(* Logix 5000 project; controller FV vendor 1 type 14 code 217 rev 31.11; software revision 31.00; part 46 of 63 *)
(* tags used below, declared in another part *)
   CWD : CHECKWORD_FLAGS;
   Delphi_Does_Eng_Func : BOOL;
   FV_FV10C : PlantItem;   // FV10C
   FV_FV10J : PlantItem;   // FV10J
   FV_FV11C : PlantItem;   // FV11C
   FV_FV11J : PlantItem;   // FV11J
   FV_FV12C : PlantItem;   // FV12C
   FV_FV12J : PlantItem;   // FV12J
   FV_FV1C : PlantItem;   // FV1C
   FV_FV1J : PlantItem;   // FV1J
   FV_FV2C : PlantItem;   // FV2C
   FV_FV2J : PlantItem;   // FV2J
   FV_FV3C : PlantItem;   // FV3C
   FV_FV3J : PlantItem;   // FV3J
   FV_FV4C : PlantItem;   // FV4C
   FV_FV4J : PlantItem;   // FV4J
   FV_FV5C : PlantItem;   // FV5C
   FV_FV5J : PlantItem;   // FV5J
   FV_FV6C : PlantItem;   // FV6C
   FV_FV6J : PlantItem;   // FV6J
   FV_FV7C : PlantItem;   // FV7C
   FV_FV7J : PlantItem;   // FV7J
   FV_FV8C : PlantItem;   // FV8C
   FV_FV8J : PlantItem;   // FV8J
   FV_FV9C : PlantItem;   // FV9C
   FV_FV9J : PlantItem;   // FV9J
   FV_N255 : INT[255];   // Old Checkwords to keep Delphi working in the interim before full changeover.
(* FV_Common, continued *)

ROUTINE FV_Old_Checkword_Relaying   (* ladder *)
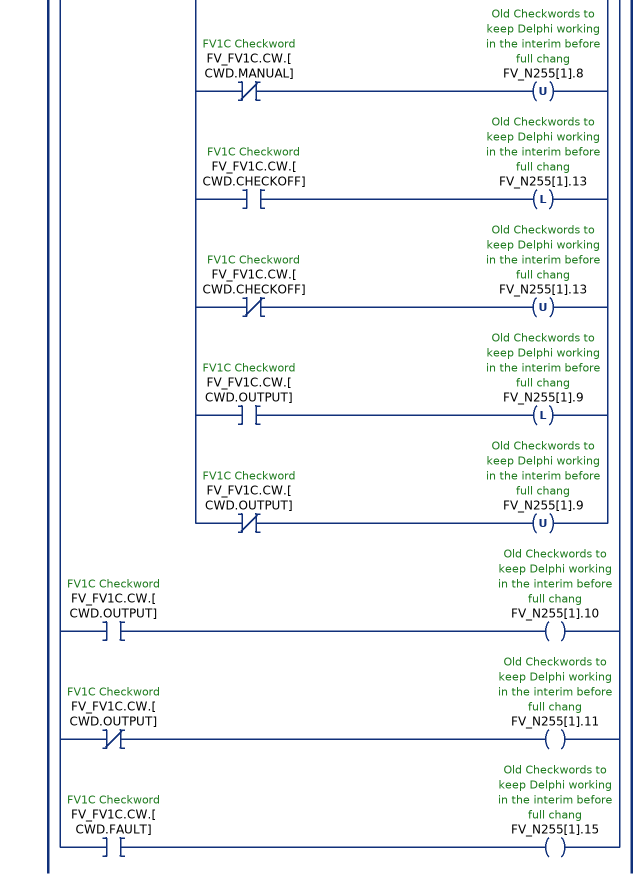
   0: [XIC(Delphi_Does_Eng_Func) [[XIC(FV_N255[1].8) [OTL(FV_FV1C.CW.[CWD.MANUAL]) ,XIC(FV_N255[1].9) OTL(FV_FV1C.CW.[CWD.MANDRV]) ,XIO(FV_N255[1].9) OTU(FV_FV1C.CW.[CWD.MANDRV]) ] ,XIO(FV_N255[1].8) [OTU(FV_FV1C.CW.[CWD.MANUAL]) ,[XIC(FV_FV1C.CW.[CWD.OUTPUT]) OTL(FV_N255[1].9) ,XIO(FV_FV1C.CW.[CWD.OUTPUT]) OTU(FV_N255[1].9) ] ] ] ,[XIC(FV_N255[1].13) OTL(FV_FV1C.CW.[CWD.CHECKOFF]) ,XIO(FV_N255[1].13) OTU(FV_FV1C.CW.[CWD.CHECKOFF]) ] ] ,XIO(Delphi_Does_Eng_Func) [[XIC(FV_FV1C.CW.[CWD.MANUAL]) OTL(FV_N255[1].8) ,XIO(FV_FV1C.CW.[CWD.MANUAL]) OTU(FV_N255[1].8) ] ,[XIC(FV_FV1C.CW.[CWD.CHECKOFF]) OTL(FV_N255[1].13) ,XIO(FV_FV1C.CW.[CWD.CHECKOFF]) OTU(FV_N255[1].13) ] ,[XIC(FV_FV1C.CW.[CWD.OUTPUT]) OTL(FV_N255[1].9) ,XIO(FV_FV1C.CW.[CWD.OUTPUT]) OTU(FV_N255[1].9) ] ] ,XIC(FV_FV1C.CW.[CWD.OUTPUT]) OTE(FV_N255[1].10) ,XIO(FV_FV1C.CW.[CWD.OUTPUT]) OTE(FV_N255[1].11) ,XIC(FV_FV1C.CW.[CWD.FAULT]) OTE(FV_N255[1].15) ];
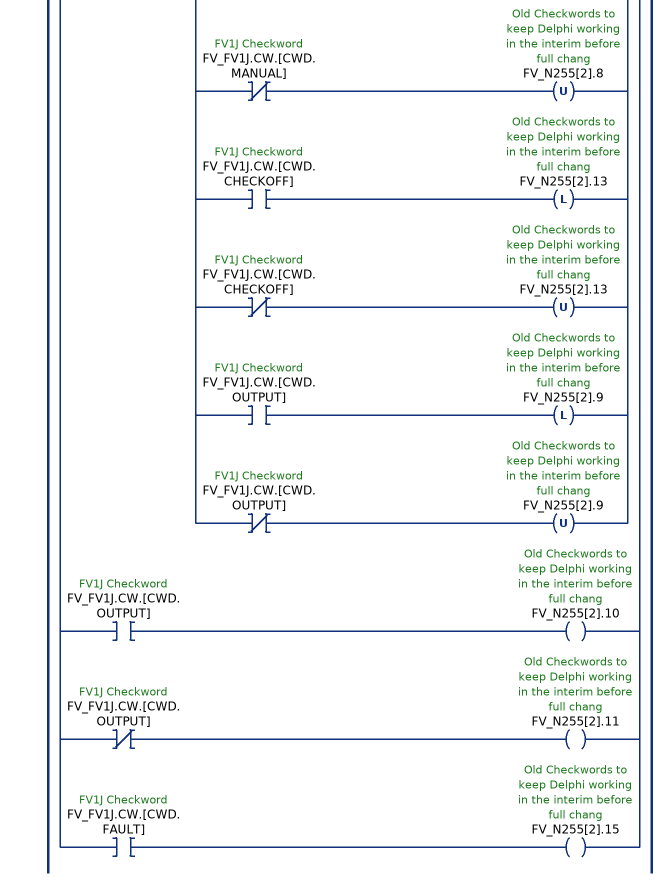
   1: [XIC(Delphi_Does_Eng_Func) [[XIC(FV_N255[2].8) [OTL(FV_FV1J.CW.[CWD.MANUAL]) ,XIC(FV_N255[2].9) OTL(FV_FV1J.CW.[CWD.MANDRV]) ,XIO(FV_N255[2].9) OTU(FV_FV1J.CW.[CWD.MANDRV]) ] ,XIO(FV_N255[2].8) [OTU(FV_FV1J.CW.[CWD.MANUAL]) ,[XIC(FV_FV1J.CW.[CWD.OUTPUT]) OTL(FV_N255[2].9) ,XIO(FV_FV1J.CW.[CWD.OUTPUT]) OTU(FV_N255[2].9) ] ] ] ,[XIC(FV_N255[2].13) OTL(FV_FV1J.CW.[CWD.CHECKOFF]) ,XIO(FV_N255[2].13) OTU(FV_FV1J.CW.[CWD.CHECKOFF]) ] ] ,XIO(Delphi_Does_Eng_Func) [[XIC(FV_FV1J.CW.[CWD.MANUAL]) OTL(FV_N255[2].8) ,XIO(FV_FV1J.CW.[CWD.MANUAL]) OTU(FV_N255[2].8) ] ,[XIC(FV_FV1J.CW.[CWD.CHECKOFF]) OTL(FV_N255[2].13) ,XIO(FV_FV1J.CW.[CWD.CHECKOFF]) OTU(FV_N255[2].13) ] ,[XIC(FV_FV1J.CW.[CWD.OUTPUT]) OTL(FV_N255[2].9) ,XIO(FV_FV1J.CW.[CWD.OUTPUT]) OTU(FV_N255[2].9) ] ] ,XIC(FV_FV1J.CW.[CWD.OUTPUT]) OTE(FV_N255[2].10) ,XIO(FV_FV1J.CW.[CWD.OUTPUT]) OTE(FV_N255[2].11) ,XIC(FV_FV1J.CW.[CWD.FAULT]) OTE(FV_N255[2].15) ];
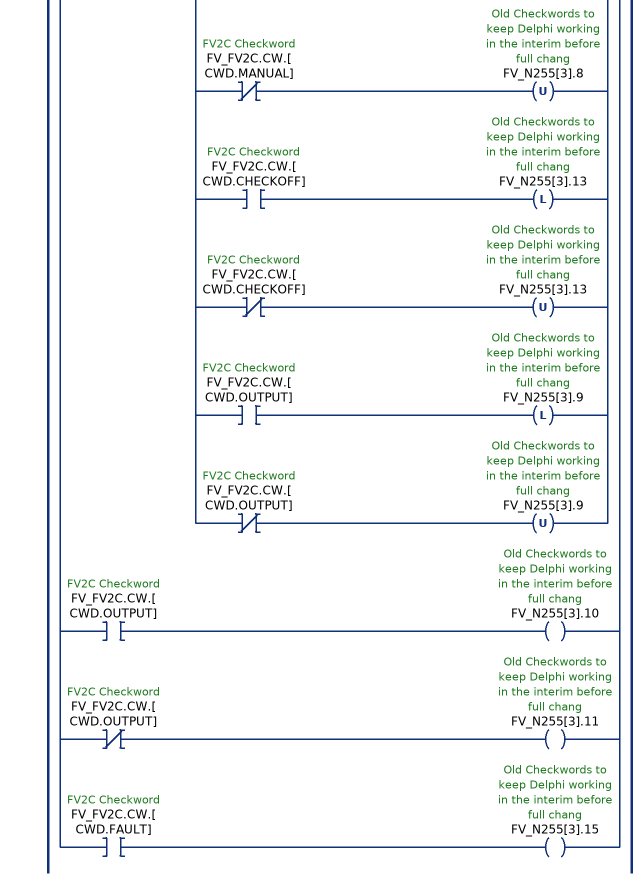
   2: [XIC(Delphi_Does_Eng_Func) [[XIC(FV_N255[3].8) [OTL(FV_FV2C.CW.[CWD.MANUAL]) ,XIC(FV_N255[3].9) OTL(FV_FV2C.CW.[CWD.MANDRV]) ,XIO(FV_N255[3].9) OTU(FV_FV2C.CW.[CWD.MANDRV]) ] ,XIO(FV_N255[3].8) [OTU(FV_FV2C.CW.[CWD.MANUAL]) ,[XIC(FV_FV2C.CW.[CWD.OUTPUT]) OTL(FV_N255[3].9) ,XIO(FV_FV2C.CW.[CWD.OUTPUT]) OTU(FV_N255[3].9) ] ] ] ,[XIC(FV_N255[3].13) OTL(FV_FV2C.CW.[CWD.CHECKOFF]) ,XIO(FV_N255[3].13) OTU(FV_FV2C.CW.[CWD.CHECKOFF]) ] ] ,XIO(Delphi_Does_Eng_Func) [[XIC(FV_FV2C.CW.[CWD.MANUAL]) OTL(FV_N255[3].8) ,XIO(FV_FV2C.CW.[CWD.MANUAL]) OTU(FV_N255[3].8) ] ,[XIC(FV_FV2C.CW.[CWD.CHECKOFF]) OTL(FV_N255[3].13) ,XIO(FV_FV2C.CW.[CWD.CHECKOFF]) OTU(FV_N255[3].13) ] ,[XIC(FV_FV2C.CW.[CWD.OUTPUT]) OTL(FV_N255[3].9) ,XIO(FV_FV2C.CW.[CWD.OUTPUT]) OTU(FV_N255[3].9) ] ] ,XIC(FV_FV2C.CW.[CWD.OUTPUT]) OTE(FV_N255[3].10) ,XIO(FV_FV2C.CW.[CWD.OUTPUT]) OTE(FV_N255[3].11) ,XIC(FV_FV2C.CW.[CWD.FAULT]) OTE(FV_N255[3].15) ];
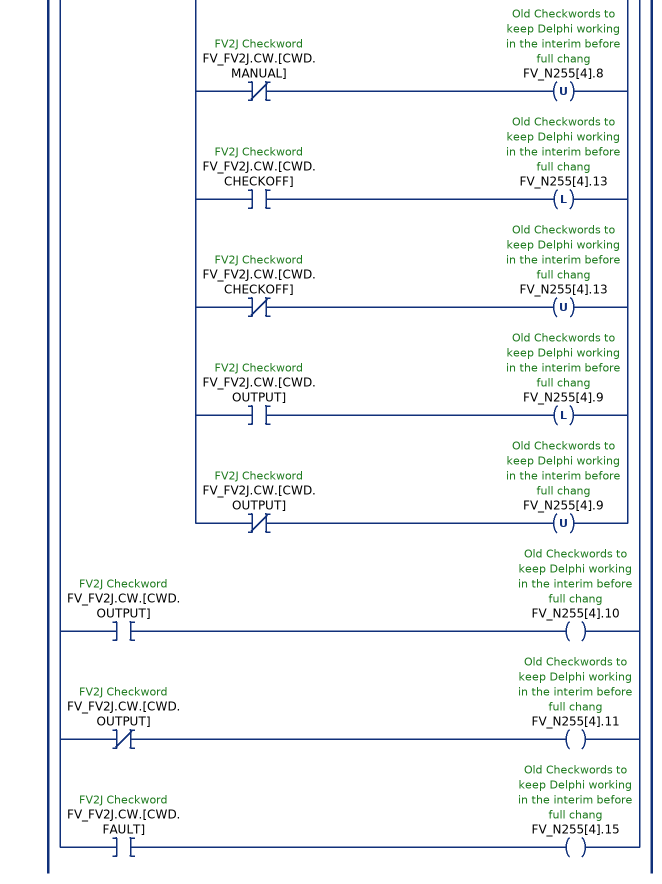
   3: [XIC(Delphi_Does_Eng_Func) [[XIC(FV_N255[4].8) [OTL(FV_FV2J.CW.[CWD.MANUAL]) ,XIC(FV_N255[4].9) OTL(FV_FV2J.CW.[CWD.MANDRV]) ,XIO(FV_N255[4].9) OTU(FV_FV2J.CW.[CWD.MANDRV]) ] ,XIO(FV_N255[4].8) [OTU(FV_FV2J.CW.[CWD.MANUAL]) ,[XIC(FV_FV2J.CW.[CWD.OUTPUT]) OTL(FV_N255[4].9) ,XIO(FV_FV2J.CW.[CWD.OUTPUT]) OTU(FV_N255[4].9) ] ] ] ,[XIC(FV_N255[4].13) OTL(FV_FV2J.CW.[CWD.CHECKOFF]) ,XIO(FV_N255[4].13) OTU(FV_FV2J.CW.[CWD.CHECKOFF]) ] ] ,XIO(Delphi_Does_Eng_Func) [[XIC(FV_FV2J.CW.[CWD.MANUAL]) OTL(FV_N255[4].8) ,XIO(FV_FV2J.CW.[CWD.MANUAL]) OTU(FV_N255[4].8) ] ,[XIC(FV_FV2J.CW.[CWD.CHECKOFF]) OTL(FV_N255[4].13) ,XIO(FV_FV2J.CW.[CWD.CHECKOFF]) OTU(FV_N255[4].13) ] ,[XIC(FV_FV2J.CW.[CWD.OUTPUT]) OTL(FV_N255[4].9) ,XIO(FV_FV2J.CW.[CWD.OUTPUT]) OTU(FV_N255[4].9) ] ] ,XIC(FV_FV2J.CW.[CWD.OUTPUT]) OTE(FV_N255[4].10) ,XIO(FV_FV2J.CW.[CWD.OUTPUT]) OTE(FV_N255[4].11) ,XIC(FV_FV2J.CW.[CWD.FAULT]) OTE(FV_N255[4].15) ];
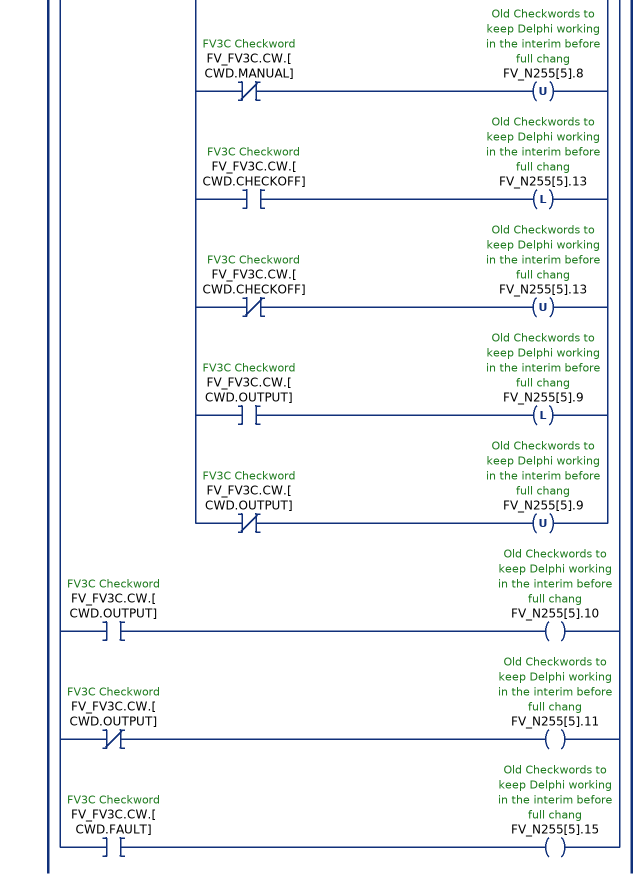
   4: [XIC(Delphi_Does_Eng_Func) [[XIC(FV_N255[5].8) [OTL(FV_FV3C.CW.[CWD.MANUAL]) ,XIC(FV_N255[5].9) OTL(FV_FV3C.CW.[CWD.MANDRV]) ,XIO(FV_N255[5].9) OTU(FV_FV3C.CW.[CWD.MANDRV]) ] ,XIO(FV_N255[5].8) [OTU(FV_FV3C.CW.[CWD.MANUAL]) ,[XIC(FV_FV3C.CW.[CWD.OUTPUT]) OTL(FV_N255[5].9) ,XIO(FV_FV3C.CW.[CWD.OUTPUT]) OTU(FV_N255[5].9) ] ] ] ,[XIC(FV_N255[5].13) OTL(FV_FV3C.CW.[CWD.CHECKOFF]) ,XIO(FV_N255[5].13) OTU(FV_FV3C.CW.[CWD.CHECKOFF]) ] ] ,XIO(Delphi_Does_Eng_Func) [[XIC(FV_FV3C.CW.[CWD.MANUAL]) OTL(FV_N255[5].8) ,XIO(FV_FV3C.CW.[CWD.MANUAL]) OTU(FV_N255[5].8) ] ,[XIC(FV_FV3C.CW.[CWD.CHECKOFF]) OTL(FV_N255[5].13) ,XIO(FV_FV3C.CW.[CWD.CHECKOFF]) OTU(FV_N255[5].13) ] ,[XIC(FV_FV3C.CW.[CWD.OUTPUT]) OTL(FV_N255[5].9) ,XIO(FV_FV3C.CW.[CWD.OUTPUT]) OTU(FV_N255[5].9) ] ] ,XIC(FV_FV3C.CW.[CWD.OUTPUT]) OTE(FV_N255[5].10) ,XIO(FV_FV3C.CW.[CWD.OUTPUT]) OTE(FV_N255[5].11) ,XIC(FV_FV3C.CW.[CWD.FAULT]) OTE(FV_N255[5].15) ];
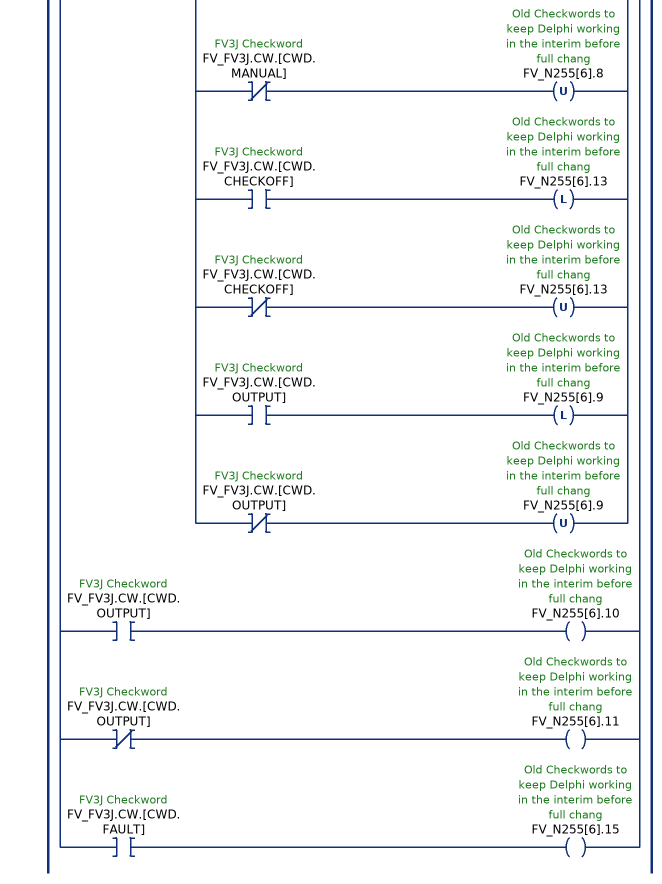
   5: [XIC(Delphi_Does_Eng_Func) [[XIC(FV_N255[6].8) [OTL(FV_FV3J.CW.[CWD.MANUAL]) ,XIC(FV_N255[6].9) OTL(FV_FV3J.CW.[CWD.MANDRV]) ,XIO(FV_N255[6].9) OTU(FV_FV3J.CW.[CWD.MANDRV]) ] ,XIO(FV_N255[6].8) [OTU(FV_FV3J.CW.[CWD.MANUAL]) ,[XIC(FV_FV3J.CW.[CWD.OUTPUT]) OTL(FV_N255[6].9) ,XIO(FV_FV3J.CW.[CWD.OUTPUT]) OTU(FV_N255[6].9) ] ] ] ,[XIC(FV_N255[6].13) OTL(FV_FV3J.CW.[CWD.CHECKOFF]) ,XIO(FV_N255[6].13) OTU(FV_FV3J.CW.[CWD.CHECKOFF]) ] ] ,XIO(Delphi_Does_Eng_Func) [[XIC(FV_FV3J.CW.[CWD.MANUAL]) OTL(FV_N255[6].8) ,XIO(FV_FV3J.CW.[CWD.MANUAL]) OTU(FV_N255[6].8) ] ,[XIC(FV_FV3J.CW.[CWD.CHECKOFF]) OTL(FV_N255[6].13) ,XIO(FV_FV3J.CW.[CWD.CHECKOFF]) OTU(FV_N255[6].13) ] ,[XIC(FV_FV3J.CW.[CWD.OUTPUT]) OTL(FV_N255[6].9) ,XIO(FV_FV3J.CW.[CWD.OUTPUT]) OTU(FV_N255[6].9) ] ] ,XIC(FV_FV3J.CW.[CWD.OUTPUT]) OTE(FV_N255[6].10) ,XIO(FV_FV3J.CW.[CWD.OUTPUT]) OTE(FV_N255[6].11) ,XIC(FV_FV3J.CW.[CWD.FAULT]) OTE(FV_N255[6].15) ];
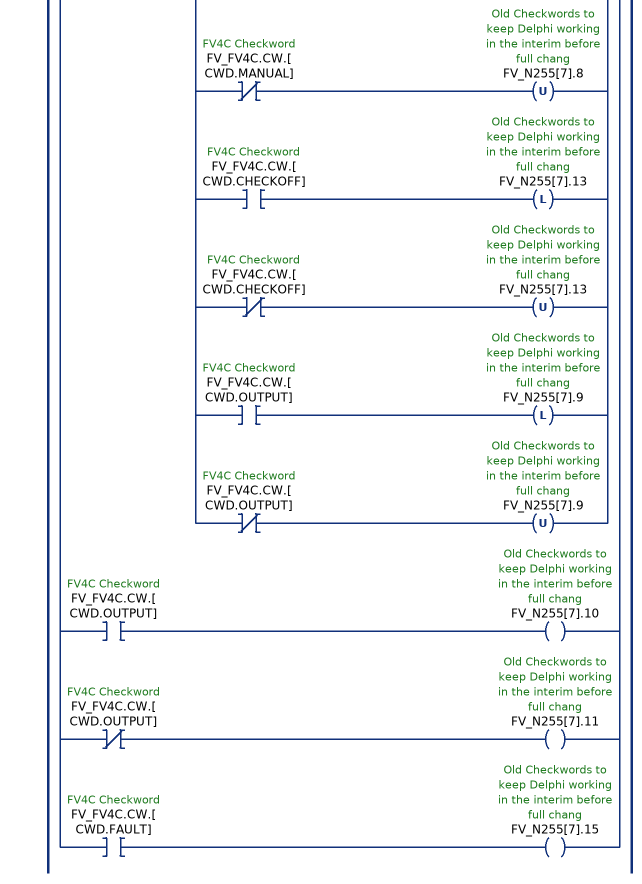
   6: [XIC(Delphi_Does_Eng_Func) [[XIC(FV_N255[7].8) [OTL(FV_FV4C.CW.[CWD.MANUAL]) ,XIC(FV_N255[7].9) OTL(FV_FV4C.CW.[CWD.MANDRV]) ,XIO(FV_N255[7].9) OTU(FV_FV4C.CW.[CWD.MANDRV]) ] ,XIO(FV_N255[7].8) [OTU(FV_FV4C.CW.[CWD.MANUAL]) ,[XIC(FV_FV4C.CW.[CWD.OUTPUT]) OTL(FV_N255[7].9) ,XIO(FV_FV4C.CW.[CWD.OUTPUT]) OTU(FV_N255[7].9) ] ] ] ,[XIC(FV_N255[7].13) OTL(FV_FV4C.CW.[CWD.CHECKOFF]) ,XIO(FV_N255[7].13) OTU(FV_FV4C.CW.[CWD.CHECKOFF]) ] ] ,XIO(Delphi_Does_Eng_Func) [[XIC(FV_FV4C.CW.[CWD.MANUAL]) OTL(FV_N255[7].8) ,XIO(FV_FV4C.CW.[CWD.MANUAL]) OTU(FV_N255[7].8) ] ,[XIC(FV_FV4C.CW.[CWD.CHECKOFF]) OTL(FV_N255[7].13) ,XIO(FV_FV4C.CW.[CWD.CHECKOFF]) OTU(FV_N255[7].13) ] ,[XIC(FV_FV4C.CW.[CWD.OUTPUT]) OTL(FV_N255[7].9) ,XIO(FV_FV4C.CW.[CWD.OUTPUT]) OTU(FV_N255[7].9) ] ] ,XIC(FV_FV4C.CW.[CWD.OUTPUT]) OTE(FV_N255[7].10) ,XIO(FV_FV4C.CW.[CWD.OUTPUT]) OTE(FV_N255[7].11) ,XIC(FV_FV4C.CW.[CWD.FAULT]) OTE(FV_N255[7].15) ];
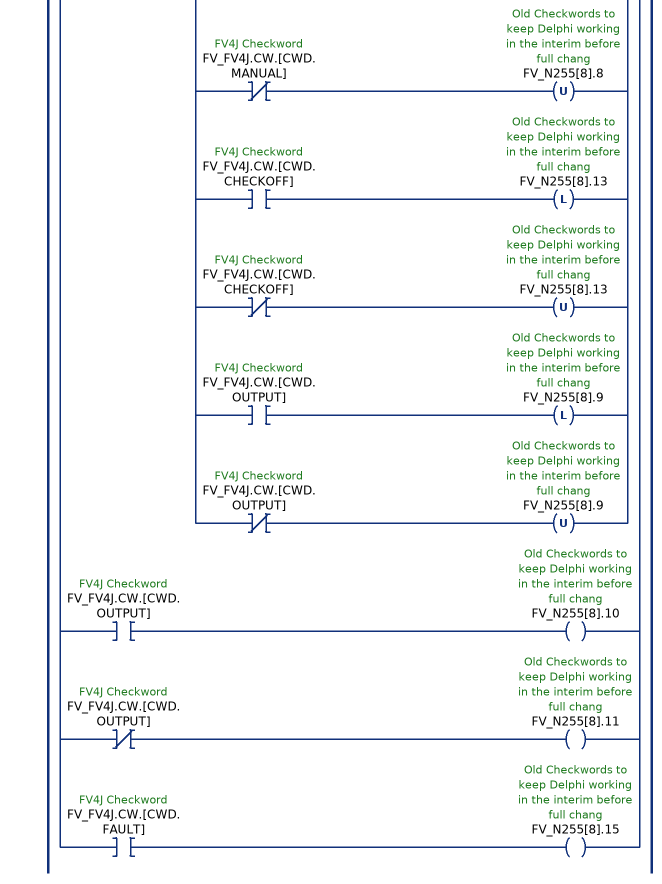
   7: [XIC(Delphi_Does_Eng_Func) [[XIC(FV_N255[8].8) [OTL(FV_FV4J.CW.[CWD.MANUAL]) ,XIC(FV_N255[8].9) OTL(FV_FV4J.CW.[CWD.MANDRV]) ,XIO(FV_N255[8].9) OTU(FV_FV4J.CW.[CWD.MANDRV]) ] ,XIO(FV_N255[8].8) [OTU(FV_FV4J.CW.[CWD.MANUAL]) ,[XIC(FV_FV4J.CW.[CWD.OUTPUT]) OTL(FV_N255[8].9) ,XIO(FV_FV4J.CW.[CWD.OUTPUT]) OTU(FV_N255[8].9) ] ] ] ,[XIC(FV_N255[8].13) OTL(FV_FV4J.CW.[CWD.CHECKOFF]) ,XIO(FV_N255[8].13) OTU(FV_FV4J.CW.[CWD.CHECKOFF]) ] ] ,XIO(Delphi_Does_Eng_Func) [[XIC(FV_FV4J.CW.[CWD.MANUAL]) OTL(FV_N255[8].8) ,XIO(FV_FV4J.CW.[CWD.MANUAL]) OTU(FV_N255[8].8) ] ,[XIC(FV_FV4J.CW.[CWD.CHECKOFF]) OTL(FV_N255[8].13) ,XIO(FV_FV4J.CW.[CWD.CHECKOFF]) OTU(FV_N255[8].13) ] ,[XIC(FV_FV4J.CW.[CWD.OUTPUT]) OTL(FV_N255[8].9) ,XIO(FV_FV4J.CW.[CWD.OUTPUT]) OTU(FV_N255[8].9) ] ] ,XIC(FV_FV4J.CW.[CWD.OUTPUT]) OTE(FV_N255[8].10) ,XIO(FV_FV4J.CW.[CWD.OUTPUT]) OTE(FV_N255[8].11) ,XIC(FV_FV4J.CW.[CWD.FAULT]) OTE(FV_N255[8].15) ];
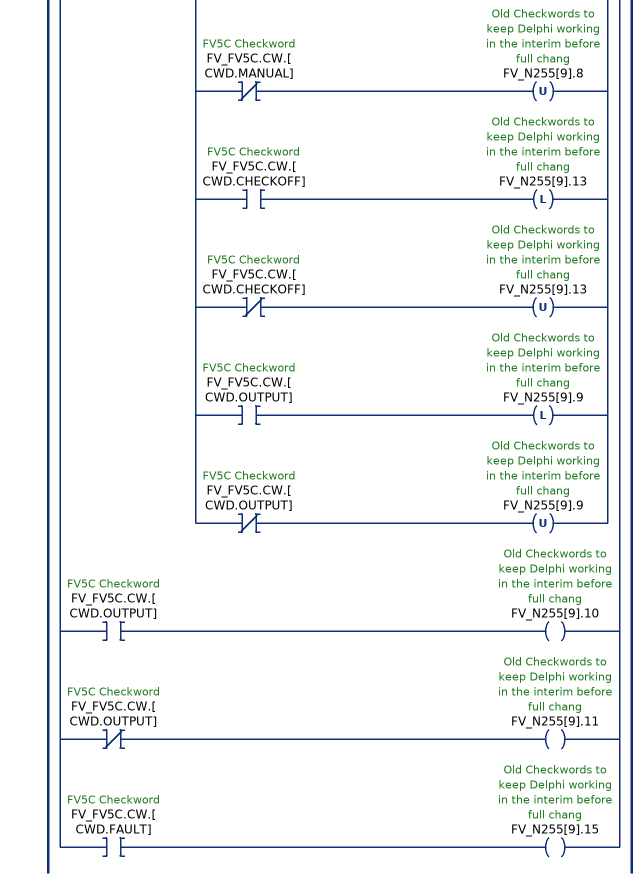
   8: [XIC(Delphi_Does_Eng_Func) [[XIC(FV_N255[9].8) [OTL(FV_FV5C.CW.[CWD.MANUAL]) ,XIC(FV_N255[9].9) OTL(FV_FV5C.CW.[CWD.MANDRV]) ,XIO(FV_N255[9].9) OTU(FV_FV5C.CW.[CWD.MANDRV]) ] ,XIO(FV_N255[9].8) [OTU(FV_FV5C.CW.[CWD.MANUAL]) ,[XIC(FV_FV5C.CW.[CWD.OUTPUT]) OTL(FV_N255[9].9) ,XIO(FV_FV5C.CW.[CWD.OUTPUT]) OTU(FV_N255[9].9) ] ] ] ,[XIC(FV_N255[9].13) OTL(FV_FV5C.CW.[CWD.CHECKOFF]) ,XIO(FV_N255[9].13) OTU(FV_FV5C.CW.[CWD.CHECKOFF]) ] ] ,XIO(Delphi_Does_Eng_Func) [[XIC(FV_FV5C.CW.[CWD.MANUAL]) OTL(FV_N255[9].8) ,XIO(FV_FV5C.CW.[CWD.MANUAL]) OTU(FV_N255[9].8) ] ,[XIC(FV_FV5C.CW.[CWD.CHECKOFF]) OTL(FV_N255[9].13) ,XIO(FV_FV5C.CW.[CWD.CHECKOFF]) OTU(FV_N255[9].13) ] ,[XIC(FV_FV5C.CW.[CWD.OUTPUT]) OTL(FV_N255[9].9) ,XIO(FV_FV5C.CW.[CWD.OUTPUT]) OTU(FV_N255[9].9) ] ] ,XIC(FV_FV5C.CW.[CWD.OUTPUT]) OTE(FV_N255[9].10) ,XIO(FV_FV5C.CW.[CWD.OUTPUT]) OTE(FV_N255[9].11) ,XIC(FV_FV5C.CW.[CWD.FAULT]) OTE(FV_N255[9].15) ];
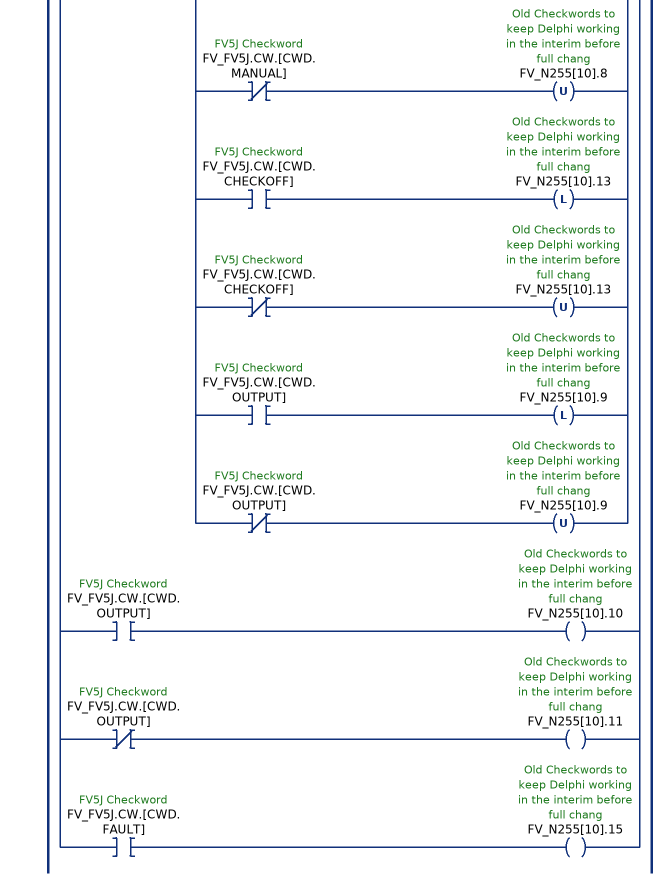
   9: [XIC(Delphi_Does_Eng_Func) [[XIC(FV_N255[10].8) [OTL(FV_FV5J.CW.[CWD.MANUAL]) ,XIC(FV_N255[10].9) OTL(FV_FV5J.CW.[CWD.MANDRV]) ,XIO(FV_N255[10].9) OTU(FV_FV5J.CW.[CWD.MANDRV]) ] ,XIO(FV_N255[10].8) [OTU(FV_FV5J.CW.[CWD.MANUAL]) ,[XIC(FV_FV5J.CW.[CWD.OUTPUT]) OTL(FV_N255[10].9) ,XIO(FV_FV5J.CW.[CWD.OUTPUT]) OTU(FV_N255[10].9) ] ] ] ,[XIC(FV_N255[10].13) OTL(FV_FV5J.CW.[CWD.CHECKOFF]) ,XIO(FV_N255[10].13) OTU(FV_FV5J.CW.[CWD.CHECKOFF]) ] ] ,XIO(Delphi_Does_Eng_Func) [[XIC(FV_FV5J.CW.[CWD.MANUAL]) OTL(FV_N255[10].8) ,XIO(FV_FV5J.CW.[CWD.MANUAL]) OTU(FV_N255[10].8) ] ,[XIC(FV_FV5J.CW.[CWD.CHECKOFF]) OTL(FV_N255[10].13) ,XIO(FV_FV5J.CW.[CWD.CHECKOFF]) OTU(FV_N255[10].13) ] ,[XIC(FV_FV5J.CW.[CWD.OUTPUT]) OTL(FV_N255[10].9) ,XIO(FV_FV5J.CW.[CWD.OUTPUT]) OTU(FV_N255[10].9) ] ] ,XIC(FV_FV5J.CW.[CWD.OUTPUT]) OTE(FV_N255[10].10) ,XIO(FV_FV5J.CW.[CWD.OUTPUT]) OTE(FV_N255[10].11) ,XIC(FV_FV5J.CW.[CWD.FAULT]) OTE(FV_N255[10].15) ];
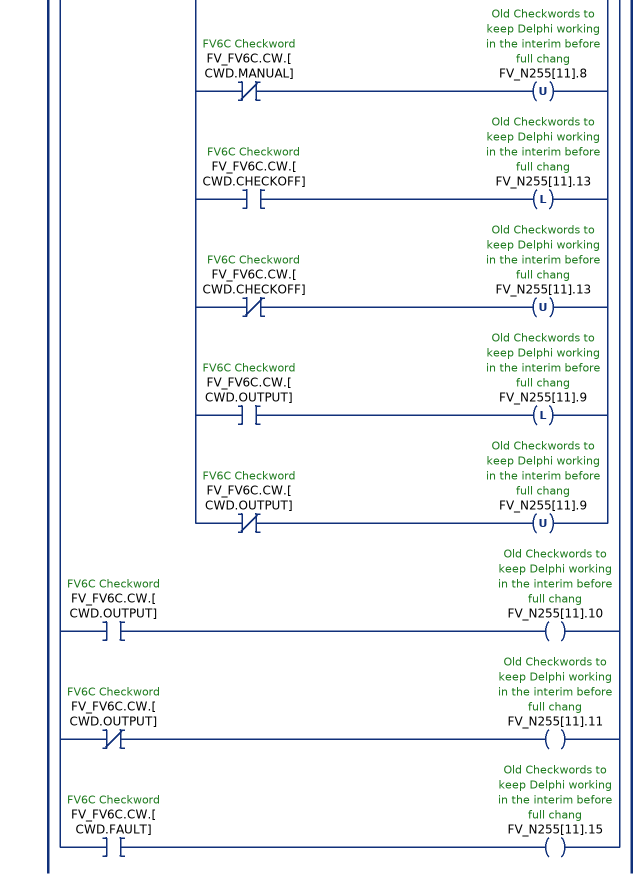
   10: [XIC(Delphi_Does_Eng_Func) [[XIC(FV_N255[11].8) [OTL(FV_FV6C.CW.[CWD.MANUAL]) ,XIC(FV_N255[11].9) OTL(FV_FV6C.CW.[CWD.MANDRV]) ,XIO(FV_N255[11].9) OTU(FV_FV6C.CW.[CWD.MANDRV]) ] ,XIO(FV_N255[11].8) [OTU(FV_FV6C.CW.[CWD.MANUAL]) ,[XIC(FV_FV6C.CW.[CWD.OUTPUT]) OTL(FV_N255[11].9) ,XIO(FV_FV6C.CW.[CWD.OUTPUT]) OTU(FV_N255[11].9) ] ] ] ,[XIC(FV_N255[11].13) OTL(FV_FV6C.CW.[CWD.CHECKOFF]) ,XIO(FV_N255[11].13) OTU(FV_FV6C.CW.[CWD.CHECKOFF]) ] ] ,XIO(Delphi_Does_Eng_Func) [[XIC(FV_FV6C.CW.[CWD.MANUAL]) OTL(FV_N255[11].8) ,XIO(FV_FV6C.CW.[CWD.MANUAL]) OTU(FV_N255[11].8) ] ,[XIC(FV_FV6C.CW.[CWD.CHECKOFF]) OTL(FV_N255[11].13) ,XIO(FV_FV6C.CW.[CWD.CHECKOFF]) OTU(FV_N255[11].13) ] ,[XIC(FV_FV6C.CW.[CWD.OUTPUT]) OTL(FV_N255[11].9) ,XIO(FV_FV6C.CW.[CWD.OUTPUT]) OTU(FV_N255[11].9) ] ] ,XIC(FV_FV6C.CW.[CWD.OUTPUT]) OTE(FV_N255[11].10) ,XIO(FV_FV6C.CW.[CWD.OUTPUT]) OTE(FV_N255[11].11) ,XIC(FV_FV6C.CW.[CWD.FAULT]) OTE(FV_N255[11].15) ];
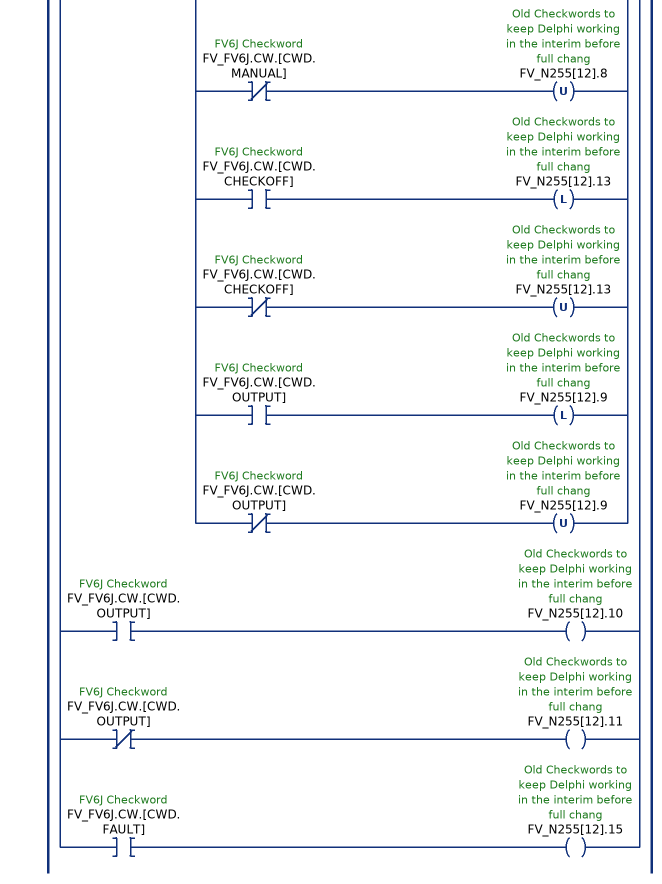
   11: [XIC(Delphi_Does_Eng_Func) [[XIC(FV_N255[12].8) [OTL(FV_FV6J.CW.[CWD.MANUAL]) ,XIC(FV_N255[12].9) OTL(FV_FV6J.CW.[CWD.MANDRV]) ,XIO(FV_N255[12].9) OTU(FV_FV6J.CW.[CWD.MANDRV]) ] ,XIO(FV_N255[12].8) [OTU(FV_FV6J.CW.[CWD.MANUAL]) ,[XIC(FV_FV6J.CW.[CWD.OUTPUT]) OTL(FV_N255[12].9) ,XIO(FV_FV6J.CW.[CWD.OUTPUT]) OTU(FV_N255[12].9) ] ] ] ,[XIC(FV_N255[12].13) OTL(FV_FV6J.CW.[CWD.CHECKOFF]) ,XIO(FV_N255[12].13) OTU(FV_FV6J.CW.[CWD.CHECKOFF]) ] ] ,XIO(Delphi_Does_Eng_Func) [[XIC(FV_FV6J.CW.[CWD.MANUAL]) OTL(FV_N255[12].8) ,XIO(FV_FV6J.CW.[CWD.MANUAL]) OTU(FV_N255[12].8) ] ,[XIC(FV_FV6J.CW.[CWD.CHECKOFF]) OTL(FV_N255[12].13) ,XIO(FV_FV6J.CW.[CWD.CHECKOFF]) OTU(FV_N255[12].13) ] ,[XIC(FV_FV6J.CW.[CWD.OUTPUT]) OTL(FV_N255[12].9) ,XIO(FV_FV6J.CW.[CWD.OUTPUT]) OTU(FV_N255[12].9) ] ] ,XIC(FV_FV6J.CW.[CWD.OUTPUT]) OTE(FV_N255[12].10) ,XIO(FV_FV6J.CW.[CWD.OUTPUT]) OTE(FV_N255[12].11) ,XIC(FV_FV6J.CW.[CWD.FAULT]) OTE(FV_N255[12].15) ];